FUNCTION_BLOCK "R-401_SEQ"   // FB30, GRAPH_PLUS
TITLE = Reactor R-401
{ S7_Optimized_Access := 'TRUE' }
AUTHOR : JL
VERSION : 0.1
   VAR_INPUT
      OFF_SQ : Bool := false;   // Turn sequence off
      INIT_SQ : Bool := false;   // Set sequence to initial state
      ACK_EF : Bool := false;   // Acknowledge all errors and faults
      S_PREV : Bool := false;   // Output previous step in parameter S_NO
      S_NEXT : Bool := false;   // Indicate next step in parameter S_NO
      SW_AUTO : Bool := false;   // Automatic mode
      SW_TAP : Bool := false;   // Semiautomatic/switch with transition
      SW_TOP : Bool := false;   // Semiautomatic/ignore transition
      SW_MAN : Bool := false;   // Manual mode
      S_SEL : Int := 0;   // Select step to be output to S_NO
      S_ON : Bool := false;   // Activate step indicated in S_NO
      S_OFF : Bool := false;   // Deactivate step indicated S_NO
      T_PUSH : Bool := false;   // Enable transition to switch in semi automatic mode
   END_VAR
   VAR_OUTPUT
      S_NO : Int := 0;   // Step number
      S_MORE : Bool := false;   // More steps are available and can be shown in S_NO
      S_ACTIVE : Bool := false;   // Step indicated in S_NO is active
      ERR_FLT : Bool := false;   // Interlock or supervision group error
      AUTO_ON : Bool := false;   // Automatic mode is active
      TAP_ON : Bool := false;   // Semiautomatic mode/step with transition enabled
      TOP_ON : Bool := false;   // Semiautomatic mode/ignore transition enabled
      MAN_ON : Bool := false;   // Manual mode is active
   END_VAR
   VAR
      HMI_INFO : Array[0..12] of UInt;
      IF_PAR : G7_IfParPlus_V6;
      RT_DATA : G7_RTDataPlus_V6;   // Internal data area
      Abort : G7_TransitionPlus_V6;   // Transition structure
      InitializeR : G7_TransitionPlus_V6;   // Transition structure
      CalcinP : G7_TransitionPlus_V6;   // Transition structure
      Re : G7_TransitionPlus_V6;   // Transition structure
      Calcinat : G7_TransitionPlus_V6;   // Transition structure
      Wash : G7_TransitionPlus_V6;   // Transition structure
      Shutdwn : G7_TransitionPlus_V6;   // Transition structure
      ColdDDn : G7_TransitionPlus_V6;   // Transition structure
      Std : G7_TransitionPlus_V6;   // Transition structure
      PDn : G7_TransitionPlus_V6;   // Transition structure
      PressRd : G7_TransitionPlus_V6;   // Transition structure
      Rmp1Dn : G7_TransitionPlus_V6;   // Transition structure
      FHldDn : G7_TransitionPlus_V6;   // Transition structure
      Rmp2Dn : G7_TransitionPlus_V6;   // Transition structure
      ScHldDn : G7_TransitionPlus_V6;   // Transition structure
      Rmp3Dn : G7_TransitionPlus_V6;   // Transition structure
      ThHldDn : G7_TransitionPlus_V6;   // Transition structure
      Trans30 : G7_TransitionPlus_V6;   // Transition structure
      Trans31 : G7_TransitionPlus_V6;   // Transition structure
      End : G7_TransitionPlus_V6;   // Transition structure
      Init : G7_TransitionPlus_V6;   // Transition structure
      SAut : G7_TransitionPlus_V6;   // Transition structure
      SIn : G7_TransitionPlus_V6;   // Transition structure
      Initd : G7_TransitionPlus_V6;   // Transition structure
      Ab : G7_TransitionPlus_V6;   // Transition structure
      AbortOn : G7_TransitionPlus_V6;   // Transition structure
      AbortDn : G7_TransitionPlus_V6;   // Transition structure
      ShtSted : G7_TransitionPlus_V6;   // Transition structure
      CldDwnDn : G7_TransitionPlus_V6;   // Transition structure
      DPDn : G7_TransitionPlus_V6;   // Transition structure
      Idle : G7_StepPlus_V6;   // Step structure
      Ready : G7_StepPlus_V6;   // Step structure
      SelectSeq : G7_StepPlus_V6;   // Step structure
      Started : G7_StepPlus_V6;   // Step structure
      "EDIT Params" : G7_StepPlus_V6;   // Step structure
      "USER StartAir" : G7_StepPlus_V6;   // Step structure
      RampUp1 : G7_StepPlus_V6;   // Step structure
      FirstHold : G7_StepPlus_V6;   // Step structure
      RampUp2 : G7_StepPlus_V6;   // Step structure
      SecondHold : G7_StepPlus_V6;   // Step structure
      RampUp3 : G7_StepPlus_V6;   // Step structure
      ThirdHold : G7_StepPlus_V6;   // Step structure
      HeatersOff : G7_StepPlus_V6;   // Step structure
      PressureOff : G7_StepPlus_V6;   // Step structure
      Done : G7_StepPlus_V6;   // Step structure
      Initialize : G7_StepPlus_V6;   // Step structure
      SetAuto : G7_StepPlus_V6;   // Step structure
      SetInitial : G7_StepPlus_V6;   // Step structure
      Initialized : G7_StepPlus_V6;   // Step structure
      AbortStarting : G7_StepPlus_V6;   // Step structure
      Aborting : G7_StepPlus_V6;   // Step structure
      AbortDone : G7_StepPlus_V6;   // Step structure
      ShtdnStarted : G7_StepPlus_V6;   // Step structure
      CoolingDown : G7_StepPlus_V6;   // Step structure
      DePress : G7_StepPlus_V6;   // Step structure
      ShtdnDn : G7_StepPlus_V6;   // Step structure
      SINI : Array[0..5] of USInt;
      LSTT : Array[0..29] of USInt;
      ATAJ : Array[0..29] of USInt;
      ATAB : Array[0..29] of USInt;
      PSTT : Array[0..29] of USInt;
      NSTT : Array[0..29] of USInt;
      ASSJ : Array[0..25] of USInt;
      ASSB : Array[0..25] of USInt;
      PTTS : Array[0..25] of USInt;
      NTTS : Array[0..25] of USInt;
      SW_SQTS : Array[0..25] of USInt;
      SWITCH : Array[0..4] of USInt;
      TVX : Array[0..11] of USInt;
      TTX : Array[0..11] of USInt;
      TSX : Array[0..5] of USInt;
      S00X : Array[0..5] of USInt;
      SOFFX : Array[0..5] of USInt;
      SONX : Array[0..5] of USInt;
      SAX : Array[0..5] of USInt;
      SERRX : Array[0..26] of USInt;
      SMX : Array[0..26] of USInt;
      S0X : Array[0..26] of USInt;
      S1X : Array[0..26] of USInt;
      IL_ALARM_INST : Diag_Alarm;
      SUP_ALARM_INST : Diag_Alarm;
      STEP_TIME_ALARM_INST : Diag_Alarm;
      IEC_TIMER_INST : IEC_TIMER;
      TRANSACTION_FLAG : Bool := false;
   END_VAR
   // SINI[0] := 2;
   // LSTT[0] := 19;
   // NSTT[0] := 19;
   // PTTS[0] := 255;
   // TVX[0] := 16#1;
   // TTX[0] := 16#1;
   // TSX[0] := 16#1;
   // S00X[0] := 16#1;
   // SOFFX[0] := 16#1;
   // SONX[0] := 16#1;
   // SAX[0] := 16#1;
   // SERRX[0] := 16#1;
   // SMX[0] := 16#1;
   // S0X[0] := 16#1;
   // S1X[0] := 16#1;
   // SINI[2] := 255;
   // SINI[3] := 255;
   // SINI[4] := 255;
   // LSTT[1] := 15;
   // LSTT[2] := 255;
   // LSTT[3] := 255;
   // LSTT[4] := 3;
   // LSTT[5] := 255;
   // LSTT[6] := 22;
   // LSTT[16] := 255;
   // LSTT[8] := 255;
   // LSTT[9] := 255;
   // LSTT[10] := 255;
   // LSTT[11] := 255;
   // LSTT[12] := 255;
   // LSTT[13] := 255;
   // LSTT[14] := 255;
   // LSTT[19] := 255;
   // LSTT[22] := 255;
   // LSTT[17] := 255;
   // LSTT[25] := 255;
   // LSTT[20] := 255;
   // LSTT[21] := 255;
   // ATAJ[1] := 1;
   // ATAJ[2] := 2;
   // ATAJ[3] := 3;
   // ATAJ[4] := 4;
   // ATAJ[5] := 5;
   // ATAJ[6] := 6;
   // ATAJ[7] := 7;
   // ATAJ[8] := 8;
   // ATAJ[9] := 9;
   // ATAJ[10] := 10;
   // ATAJ[11] := 11;
   // ATAJ[12] := 12;
   // ATAJ[13] := 13;
   // ATAJ[14] := 14;
   // ATAJ[15] := 15;
   // ATAJ[16] := 16;
   // ATAJ[17] := 17;
   // ATAJ[18] := 18;
   // ATAJ[19] := 19;
   // ATAJ[20] := 20;
   // ATAJ[21] := 21;
   // ATAJ[22] := 22;
   // ATAB[0] := 6;
   // ATAB[1] := 2;
   // ATAB[3] := 3;
   // ATAB[4] := 5;
   // ATAB[5] := 4;
   // ATAB[6] := 1;
   // ATAB[7] := 7;
   // ATAB[8] := 8;
   // ATAB[9] := 9;
   // ATAB[10] := 10;
   // ATAB[11] := 11;
   // ATAB[12] := 12;
   // ATAB[13] := 13;
   // ATAB[14] := 14;
   // ATAB[15] := 15;
   // ATAB[16] := 16;
   // ATAB[17] := 17;
   // ATAB[18] := 18;
   // ATAB[19] := 19;
   // ATAB[20] := 20;
   // ATAB[21] := 21;
   // ATAB[22] := 22;
   // SW_SQTS[21] := 4;
   // SW_SQTS[20] := 4;
   // PSTT[3] := 1;
   // PSTT[4] := 2;
   // PSTT[5] := 2;
   // PSTT[22] := 17;
   // PSTT[7] := 25;
   // PSTT[8] := 3;
   // PSTT[9] := 4;
   // PSTT[10] := 5;
   // PSTT[11] := 6;
   // PSTT[12] := 7;
   // PSTT[13] := 8;
   // PSTT[14] := 9;
   // PSTT[15] := 10;
   // PSTT[16] := 11;
   // PSTT[17] := 13;
   // PSTT[18] := 14;
   // PSTT[19] := 12;
   // PSTT[20] := 15;
   // PSTT[21] := 16;
   // PSTT[25] := 20;
   // NTTS[21] := 26;
   // NTTS[20] := 25;
   // PTTS[21] := 25;
   // PTTS[20] := 24;
   // NSTT[1] := 15;
   // NSTT[2] := 1;
   // NSTT[3] := 2;
   // NSTT[4] := 3;
   // NSTT[5] := 255;
   // NSTT[6] := 22;
   // NSTT[16] := 12;
   // NSTT[8] := 4;
   // NSTT[9] := 5;
   // NSTT[10] := 6;
   // NSTT[11] := 7;
   // NSTT[12] := 8;
   // NSTT[13] := 9;
   // NSTT[14] := 10;
   // NSTT[19] := 13;
   // NSTT[22] := 18;
   // NSTT[17] := 14;
   // NSTT[25] := 21;
   // NSTT[20] := 16;
   // NSTT[21] := 17;
   // ASSJ[20] := 20;
   // ASSB[21] := 21;
   // ASSB[20] := 20;
   // ASSJ[21] := 21;
   // ASSJ[1] := 1;
   // ASSJ[2] := 2;
   // ASSJ[3] := 3;
   // ASSJ[4] := 4;
   // ASSJ[5] := 5;
   // ASSJ[6] := 6;
   // ASSJ[7] := 7;
   // ASSJ[8] := 8;
   // ASSJ[9] := 9;
   // ASSJ[10] := 10;
   // ASSJ[11] := 11;
   // ASSJ[12] := 12;
   // ASSJ[13] := 13;
   // ASSJ[14] := 14;
   // ASSJ[15] := 15;
   // ASSJ[16] := 16;
   // ASSJ[17] := 17;
   // ASSJ[18] := 18;
   // ASSJ[19] := 19;
   // NSTT[23] := 1;
   // NSTT[15] := 11;
   // PSTT[24] := 19;
   // PSTT[23] := 18;
   // ASSB[1] := 1;
   // ASSB[2] := 2;
   // ASSB[3] := 3;
   // ASSB[4] := 4;
   // ASSB[5] := 5;
   // ASSB[6] := 6;
   // ASSB[7] := 7;
   // ASSB[8] := 8;
   // ASSB[9] := 9;
   // ASSB[10] := 10;
   // ASSB[11] := 11;
   // ASSB[12] := 12;
   // ASSB[13] := 13;
   // ASSB[14] := 14;
   // ASSB[15] := 15;
   // ASSB[16] := 16;
   // ASSB[17] := 17;
   // ASSB[18] := 18;
   // ASSB[19] := 19;
   // ATAB[24] := 24;
   // ATAB[23] := 23;
   // ATAJ[24] := 24;
   // ATAJ[23] := 23;
   // PTTS[1] := 2;
   // PTTS[2] := 3;
   // PTTS[3] := 255;
   // PTTS[4] := 8;
   // PTTS[5] := 9;
   // PTTS[6] := 10;
   // PTTS[7] := 11;
   // PTTS[8] := 12;
   // PTTS[9] := 13;
   // PTTS[10] := 14;
   // PTTS[11] := 15;
   // PTTS[12] := 16;
   // PTTS[13] := 19;
   // PTTS[14] := 17;
   // PTTS[15] := 255;
   // PTTS[16] := 20;
   // PTTS[17] := 21;
   // PTTS[18] := 22;
   // PTTS[19] := 255;
   // LSTT[23] := 1;
   // LSTT[15] := 255;
   // NTTS[1] := 3;
   // NTTS[2] := 4;
   // NTTS[3] := 8;
   // NTTS[4] := 9;
   // NTTS[5] := 10;
   // NTTS[6] := 11;
   // NTTS[7] := 12;
   // NTTS[8] := 13;
   // NTTS[9] := 14;
   // NTTS[10] := 15;
   // NTTS[11] := 16;
   // NTTS[12] := 19;
   // NTTS[13] := 17;
   // NTTS[14] := 18;
   // NTTS[15] := 20;
   // NTTS[16] := 21;
   // NTTS[17] := 22;
   // NTTS[18] := 23;
   // NTTS[19] := 24;
   // SW_SQTS[1] := 1;
   // SW_SQTS[2] := 1;
   // SW_SQTS[3] := 2;
   // SW_SQTS[4] := 2;
   // SW_SQTS[5] := 2;
   // SW_SQTS[6] := 2;
   // SW_SQTS[7] := 2;
   // SW_SQTS[8] := 2;
   // SW_SQTS[9] := 2;
   // SW_SQTS[10] := 2;
   // SW_SQTS[11] := 2;
   // SW_SQTS[12] := 2;
   // SW_SQTS[13] := 2;
   // SW_SQTS[14] := 2;
   // SW_SQTS[15] := 3;
   // SW_SQTS[16] := 3;
   // SW_SQTS[17] := 3;
   // SW_SQTS[18] := 3;
   // SW_SQTS[19] := 4;
   // SWITCH[0] := 60;
   // SWITCH[1] := 191;
   // SWITCH[2] := 223;
   // SINI[5] := 255;
   // LSTT[24] := 255;
   // LSTT[28] := 255;
   // LSTT[27] := 255;
   // ATAJ[25] := 25;
   // ATAJ[26] := 26;
   // ATAJ[27] := 27;
   // ATAJ[28] := 28;
   // ATAB[25] := 25;
   // ATAB[26] := 26;
   // ATAB[27] := 27;
   // ATAB[28] := 28;
   // PSTT[26] := 21;
   // PSTT[27] := 22;
   // PSTT[28] := 23;
   // NSTT[24] := 20;
   // NSTT[28] := 24;
   // NSTT[27] := 23;
   // ASSJ[22] := 22;
   // ASSJ[23] := 23;
   // ASSJ[24] := 24;
   // ASSB[22] := 22;
   // ASSB[23] := 23;
   // ASSB[24] := 24;
   // PTTS[22] := 255;
   // PTTS[23] := 27;
   // PTTS[24] := 28;
   // NTTS[22] := 27;
   // NTTS[23] := 28;
   // NTTS[24] := 29;
   // SW_SQTS[22] := 5;
   // SW_SQTS[23] := 5;
   // SW_SQTS[24] := 5;
   // SWITCH[3] := 239;
   // SWITCH[4] := 7;
   // LSTT[29] := 255;
   // ATAJ[29] := 29;
   // ATAB[29] := 29;
   // PSTT[29] := 24;
   // NSTT[29] := 25;
   // ASSJ[25] := 25;
   // ASSB[25] := 25;
   // PTTS[25] := 29;
   // NTTS[25] := 7;
   // SW_SQTS[25] := 5;
BEGIN
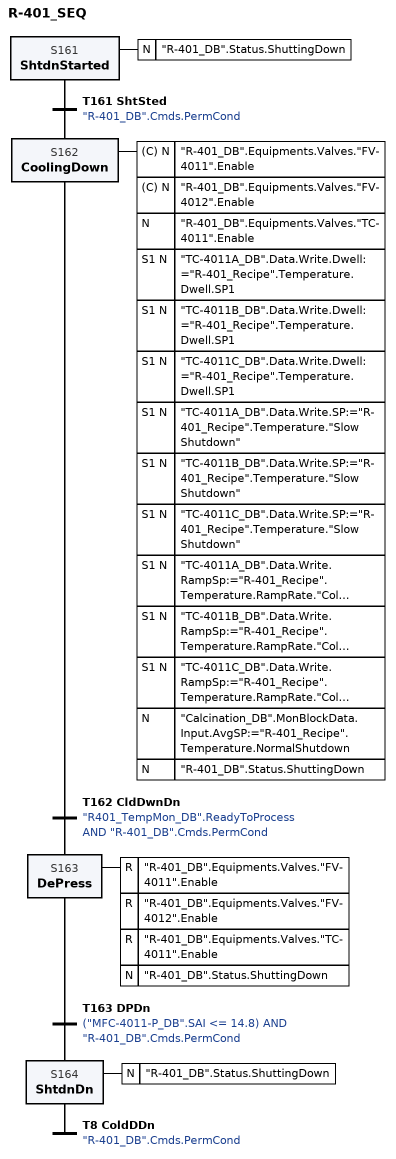
   // permanent pre-instructions
   NETWORK 1
      "R-401_SEQ_FC"();
      "R-401_FC_Inputs"();
      "Monitor_SEQ_FC"();
      "R-401_Tansitions_FC"();
      "Alarms"();

   // sequencer 1
   STEP ShtdnStarted:   // S161, max time T#10S, warning time T#7S
      // Shutdown Started
              N    "R-401_DB".Status.ShuttingDown
   END_STEP
   TRANSITION ShtSted FROM ShtdnStarted TO CoolingDown   // T161
      := "R-401_DB".Cmds.PermCond;
   END_TRANSITION
   STEP CoolingDown:   // S162, max time T#10S, warning time T#7S
      interlock C := "R-401_DB".Cmds.IL;
      (C)     N    "R-401_DB".Equipments.Valves."FV-4011".Enable
      (C)     N    "R-401_DB".Equipments.Valves."FV-4012".Enable
              N    "R-401_DB".Equipments.Valves."TC-4011".Enable
          S1  N    "TC-4011A_DB".Data.Write.Dwell:="R-401_Recipe".Temperature.Dwell.SP1
          S1  N    "TC-4011B_DB".Data.Write.Dwell:="R-401_Recipe".Temperature.Dwell.SP1
          S1  N    "TC-4011C_DB".Data.Write.Dwell:="R-401_Recipe".Temperature.Dwell.SP1
          S1  N    "TC-4011A_DB".Data.Write.SP:="R-401_Recipe".Temperature."Slow Shutdown"
          S1  N    "TC-4011B_DB".Data.Write.SP:="R-401_Recipe".Temperature."Slow Shutdown"
          S1  N    "TC-4011C_DB".Data.Write.SP:="R-401_Recipe".Temperature."Slow Shutdown"
          S1  N    "TC-4011A_DB".Data.Write.RampSp:="R-401_Recipe".Temperature.RampRate."Cold Down"
          S1  N    "TC-4011B_DB".Data.Write.RampSp:="R-401_Recipe".Temperature.RampRate."Cold Down"
          S1  N    "TC-4011C_DB".Data.Write.RampSp:="R-401_Recipe".Temperature.RampRate."Cold Down"
              N    "Calcination_DB".MonBlockData.Input.AvgSP:="R-401_Recipe".Temperature.NormalShutdown
              N    "R-401_DB".Status.ShuttingDown
   END_STEP
   TRANSITION CldDwnDn FROM CoolingDown TO DePress   // T162
      := "R401_TempMon_DB".ReadyToProcess AND "R-401_DB".Cmds.PermCond;
   END_TRANSITION
   STEP DePress:   // S163, max time T#10S, warning time T#7S
              R    "R-401_DB".Equipments.Valves."FV-4011".Enable
              R    "R-401_DB".Equipments.Valves."FV-4012".Enable
              R    "R-401_DB".Equipments.Valves."TC-4011".Enable
              N    "R-401_DB".Status.ShuttingDown
   END_STEP
   TRANSITION DPDn FROM DePress TO ShtdnDn   // T163
      := ("MFC-4011-P_DB".SAI <= 14.8) AND "R-401_DB".Cmds.PermCond;
   END_TRANSITION
   STEP ShtdnDn:   // S164, max time T#10S, warning time T#7S
              N    "R-401_DB".Status.ShuttingDown
   END_STEP
   TRANSITION ColdDDn FROM ShtdnDn TO ?   // T8
      := "R-401_DB".Cmds.PermCond;
   END_TRANSITION

   // permanent post-instructions
   NETWORK 1
      "R-401_FC_Outputs"();
END_FUNCTION_BLOCK

FUNCTION "R-401_FC_Inputs" : Void   // FC51, SCL
{ S7_Optimized_Access := 'TRUE' }
VERSION : 0.1
   VAR_TEMP
      fdfdfd : DInt;
   END_VAR
BEGIN
   //************************************************************************************************************************************
   //************************************************From Eurotherm TC-401A Controllers*********************************************************
   //***************************************************** Working Setpoint (SP)********************************************************

   IF "R-402_Aux_DB"."Bool".EurothermStatus."4011A_Connected" THEN     //Check if Modbus Connection is Ok
       "TC-4011A_DB".Data.Read.WorkingSP := INT_TO_REAL("TC-4011A_R1".MB_Data.Buffer[5]);
   ELSE
       "TC-4011A_DB".Data.Read.WorkingSP := 0.0;
   END_IF;

   IF "R-402_Aux_DB"."Bool".EurothermStatus."4011B_Connected" THEN     //Check if Modbus Connection is Ok
       "TC-4011B_DB".Data.Read.WorkingSP := INT_TO_REAL("TC-4011B_R1".MB_Data.Buffer[5]);
   ELSE
       "TC-4011B_DB".Data.Read.WorkingSP := 0.0;
   END_IF;

   IF "R-402_Aux_DB"."Bool".EurothermStatus."4011C_Connected" THEN     //Check if Modbus Connection is Ok
       "TC-4011C_DB".Data.Read.WorkingSP := INT_TO_REAL("TC-4011C_R1".MB_Data.Buffer[5]);
   ELSE
       "TC-4011C_DB".Data.Read.WorkingSP := 0.0;
   END_IF;

   //*****************************************************Process Value (PV)********************************************************

   IF "R-402_Aux_DB"."Bool".EurothermStatus."4011A_Connected" THEN     //Check if Modbus Connection is Ok
       "TC-4011A_DB".Data.Read.PV := INT_TO_REAL("TC-4011A_R1".MB_Data.Buffer[1]);
   ELSE
       "TC-4011A_DB".Data.Read.PV := 0.0;
   END_IF;

   IF "R-402_Aux_DB"."Bool".EurothermStatus."4011B_Connected" THEN     //Check if Modbus Connection is Ok
       "TC-4011B_DB".Data.Read.PV := INT_TO_REAL("TC-4011B_R1".MB_Data.Buffer[1]);
   ELSE
       "TC-4011B_DB".Data.Read.PV := 0.0;
   END_IF;

   IF "R-402_Aux_DB"."Bool".EurothermStatus."4011C_Connected" THEN     //Check if Modbus Connection is Ok
       "TC-4011C_DB".Data.Read.PV := INT_TO_REAL("TC-4011C_R1".MB_Data.Buffer[1]);
   ELSE
       "TC-4011C_DB".Data.Read.PV := 0.0;
   END_IF;


   //***************************************************** Controller Output (OP)******************************************************

   IF "R-402_Aux_DB"."Bool".EurothermStatus."4011A_Connected" THEN     //Check if Modbus Connection is Ok
       "TC-4011A_DB".Data.Read.OP := INT_TO_REAL("TC-4011A_R1".MB_Data.Buffer[4]/10);
   ELSE
       "TC-4011A_DB".Data.Read.OP := 0.0;
   END_IF;

   IF "R-402_Aux_DB"."Bool".EurothermStatus."4011B_Connected" THEN     //Check if Modbus Connection is Ok
       "TC-4011B_DB".Data.Read.OP := INT_TO_REAL("TC-4011B_R1".MB_Data.Buffer[4] / 10);
   ELSE
       "TC-4011B_DB".Data.Read.OP := 0.0;
   END_IF;

   IF "R-402_Aux_DB"."Bool".EurothermStatus."4011C_Connected" THEN     //Check if Modbus Connection is Ok
       "TC-4011C_DB".Data.Read.OP := INT_TO_REAL("TC-4011C_R1".MB_Data.Buffer[4]/10);
   ELSE
       "TC-4011C_DB".Data.Read.OP := 0.0;
   END_IF;
END_FUNCTION

FUNCTION "R-401_FC_Outputs" : Void   // FC85, SCL
{ S7_Optimized_Access := 'TRUE' }
VERSION : 0.1
   VAR_TEMP
      "FV-4011" : Struct
         On : Bool;
         Cond_1 : Bool;
      END_STRUCT;
      "FV-4012" : Struct
         On : Bool;
         Cond_1 : Bool;
      END_STRUCT;
      "TC-4011" : Struct
         On : Bool;
         Cond_1 : Bool;
      END_STRUCT;
   END_VAR
BEGIN
   //****** Equipmens Activation*******
   //**********************************TC-4011 Eurotherm Temperature Control (TC-4011)**************************************************

   #"TC-4011".Cond_1 := "R-401_DB".Equipments.Valves."TC-4011".Enable AND NOT "R-401_Aux_DB".Timer.HoldTimer.Q;
       "R-401_DB".Equipments.Valves."TC-4011".CmdOn := #"TC-4011".Cond_1 AND NOT "R-401_DB".Cmds.Hold AND NOT "R-401_DB".Status.Aborting;
       //Delay Off 
       #"TC-4011".On := "R-401_DB".Equipments.Valves."TC-4011".CmdOn;

       IF #"TC-4011".On AND ("R-401_DB".Status.Step=24 OR "R-401_DB".Status.Step=26 OR "R-401_DB".Status.Step=28) AND "R-401_Aux_DB"."Bool".Cond._005 THEN //Run Command for the Eurotherm Controllers
           "TC-4011A_DB".Data.Write.CMD := 1;
           "TC-4011B_DB".Data.Write.CMD  := 1;
           "TC-4011C_DB".Data.Write.CMD  := 1;

           //**********Working SP Reached ********
           "R-401_Aux_DB"."Bool".Cond._006 := "TC-4011A_DB".Data.Write.SP = "TC-4011A_DB".Data.Read.WorkingSP;
           "R-401_Aux_DB"."Bool".Cond._007 := "TC-4011B_DB".Data.Write.SP = "TC-4011B_DB".Data.Read.WorkingSP;
           "R-401_Aux_DB"."Bool".Cond._008 := "TC-4011C_DB".Data.Write.SP = "TC-4011C_DB".Data.Read.WorkingSP;

           "R-401_Aux_DB"."Bool".Cond._009 := "R-401_Aux_DB"."Bool".Cond._006 AND "R-401_Aux_DB"."Bool".Cond._007 AND "R-401_Aux_DB"."Bool".Cond._008;

       ELSIF #"TC-4011".On AND ("R-401_DB".Status.Step=25 OR "R-401_DB".Status.Step=27 OR "R-401_DB".Status.Step=29) AND "R-401_Aux_DB"."Bool".Cond._005 THEN //Hold command for the Eurotherm Controllers
           "TC-4011A_DB".Data.Write.CMD  := 2;
           "TC-4011B_DB".Data.Write.CMD  := 2;
           "TC-4011C_DB".Data.Write.CMD  := 2;

           "R-401_Aux_DB"."Bool".Cond._009 := FALSE;
       ELSE    //Stop Command for the Eurotherm Controllers
           "TC-4011A_DB".Data.Write.CMD  := 0;
           "TC-4011B_DB".Data.Write.CMD  := 0;
           "TC-4011C_DB".Data.Write.CMD  := 0;

           "R-401_Aux_DB"."Bool".Cond._009 := FALSE;
       END_IF;
       "R-401_DB".Equipments.Valves."TC-4011".TurningOff := NOT "R-401_DB".Equipments.Valves."TC-4011".CmdOn AND "R-401_Aux_DB".Timer."TC-4011".Q;

   //**********************************FV-4011 Air Pressure Control Valve (MFC-4011)******************************************************
   IF "FV-4011_DB".HMI.Config.Mode = 0 THEN
       #"FV-4011".Cond_1 := "R-401_DB".Equipments.Valves."FV-4011".Enable;
       "R-401_DB".Equipments.Valves."FV-4011".CmdOn := #"FV-4011".Cond_1 AND NOT "R-401_DB".Cmds.Hold AND NOT "R-401_DB".Status.Aborting;
       //Delay Off To avoid Overpressure the Lines
       #"FV-4011".On := "R-401_DB".Equipments.Valves."FV-4011".CmdOn;
       "R-401_Aux_DB".Timer."FV-4011".TOF(IN := #"FV-4011".On,
                                          PT := "R-401_Aux_DB".Constants.CmdDelay);
       IF "R-401_Aux_DB".Timer."FV-4011".Q  THEN

           // "MFC-4011_DB_MB".Data.SP := "R-401_Recipe".Pressure.Calcination;

           "MFC-4011_DB".enableManualMode := False;
           "MFC-4011_DB".enableRemoteSetpoint := False;
            "MFC-4011_DB".hmi.Controls.manualEnable := False;
            "MFC-4011_DB".hmi.Config.mode := 3;

       END_IF;
      // ELSE
          // "MFC-4011_DB".enableManualMode := True;
          // "MFC-4011_DB".hmi.Controls.manualEnable := True;
          // "MFC-4011_DB".hmi.Config.mode := 4;
          // "MFC-4011_DB".hmi.Controls.manualOutput := "R-401_Recipe".Pressure.Shutdown;

          // "MFC-4011_DB_MB".Data.SP := "R-401_Recipe".Pressure.Shutdown;

      // END_IF;
       "R-401_DB".Equipments.Valves."FV-4011".TurningOff := NOT "R-401_DB".Equipments.Valves."FV-4011".CmdOn AND "R-401_Aux_DB".Timer."FV-4011".Q;
   END_IF;

   //**********************************FV-4012 N2 Pressure Control Valve (MFC-4012)******************************************************
   IF "FV-4012_DB".HMI.Config.Mode = 0 THEN
       #"FV-4012".Cond_1 := "R-401_DB".Equipments.Valves."FV-4012".Enable;
       "R-401_DB".Equipments.Valves."FV-4012".CmdOn := #"FV-4012".Cond_1 AND NOT "R-401_DB".Cmds.Hold AND NOT "R-401_DB".Status.Aborting;
       //Delay Off To avoid Overpressure the Lines
       #"FV-4012".On := "R-401_DB".Equipments.Valves."FV-4012".CmdOn;
       "R-401_Aux_DB".Timer."FV-4012".TOF(IN := #"FV-4012".On,
                                          PT := "R-401_Aux_DB".Constants.CmdDelay);
       IF "R-401_Aux_DB".Timer."FV-4012".Q THEN

           // "MFC-4011_DB_MB".Data.SP := "R-401_Recipe".Pressure.Calcination;

           "MFC-4012_DB".enableManualMode := False;
           "MFC-4012_DB".enableRemoteSetpoint := False;
           "MFC-4012_DB".hmi.Controls.manualEnable := False;
           "MFC-4012_DB".hmi.Config.mode := 3;

       END_IF;
       // ELSE
       // "MFC-4011_DB".enableManualMode := True;
       // "MFC-4011_DB".hmi.Controls.manualEnable := True;
       // "MFC-4011_DB".hmi.Config.mode := 4;
       // "MFC-4011_DB".hmi.Controls.manualOutput := "R-401_Recipe".Pressure.Shutdown;

       // "MFC-4011_DB_MB".Data.SP := "R-401_Recipe".Pressure.Shutdown;

       // END_IF;
       "R-401_DB".Equipments.Valves."FV-4012".TurningOff := NOT "R-401_DB".Equipments.Valves."FV-4012".CmdOn AND "R-401_Aux_DB".Timer."FV-4012".Q;
   END_IF;
   //******************************************************************************************************************************************//
   //**************************************************To Temperature Controllers**************************************************************

       //***********************************************Temperature Controllers Commands*******************************************************//
   "TC-4011A_W1".MB_Data.Buffer[1] := "TC-4011A_DB".Data.Write.CMD;
   "TC-4011B_W1".MB_Data.Buffer[1]:= "TC-4011B_DB".Data.Write.CMD;
   "TC-4011C_W1".MB_Data.Buffer[1] := "TC-4011C_DB".Data.Write.CMD;

   //***********************************************Dwell to Temperature Controllers ******************************************************//
   IF "TC-4011A_DB".Data.Write.Dwell = "TC-4011A_R2".MB_Data.Buffer[1]
       AND "TC-4011A_DB".Data.Write.Dwell = "TC-4011B_R2".MB_Data.Buffer[1]
       AND "TC-4011A_DB".Data.Write.Dwell = "TC-4011C_R2".MB_Data.Buffer[1] THEN    //Compare read value and SP to activate or deactivate the Modbus Write block

       "TC-4011A_W2".Disconnect := TRUE;
       "TC-4011B_W2".Disconnect := TRUE;
       "TC-4011C_W2".Disconnect := TRUE;
       "R-401_Aux_DB"."Bool".Cond._004 := TRUE;
   ELSE
       "TC-4011A_W2".MB_Data.Buffer[1] := "TC-4011A_DB".Data.Write.Dwell;
       "TC-4011B_W2".MB_Data.Buffer[1] := "TC-4011B_DB".Data.Write.Dwell;
       "TC-4011C_W2".MB_Data.Buffer[1] := "TC-4011C_DB".Data.Write.Dwell;
       "TC-4011A_W2".Disconnect := FALSE;
       "TC-4011B_W2".Disconnect := FALSE;
       "TC-4011C_W2".Disconnect := FALSE;
       "R-401_Aux_DB"."Bool".Cond._004 := FALSE;
   END_IF;
       //***********************************************Temperature Controllers SetPoints*****************************************************//
   IF "TC-4011A_DB".Data.Write.SP = "TC-4011A_R2".MB_Data.Buffer[2]    
       AND "TC-4011A_DB".Data.Write.SP = "TC-4011B_R2".MB_Data.Buffer[2]
       AND "TC-4011A_DB".Data.Write.SP = "TC-4011C_R2".MB_Data.Buffer[2] THEN   //Compare read value and SP to activate or deactivate the Modbus Write block
       "TC-4011A_W3".Disconnect := TRUE;
       "TC-4011B_W3".Disconnect := TRUE;
       "TC-4011C_W3".Disconnect := TRUE;
       "R-401_Aux_DB"."Bool".Cond._002 := TRUE;        //Temperature SP
   ELSE
       "TC-4011A_W3".MB_Data.Buffer[1] := REAL_TO_INT("TC-4011A_DB".Data.Write.SP);
       "TC-4011B_W3".MB_Data.Buffer[1] := REAL_TO_INT("TC-4011B_DB".Data.Write.SP);
       "TC-4011C_W3".MB_Data.Buffer[1] := REAL_TO_INT("TC-4011C_DB".Data.Write.SP);
       "TC-4011A_W3".Disconnect := FALSE;
       "TC-4011B_W3".Disconnect := FALSE;
       "TC-4011C_W3".Disconnect := FALSE;
       "R-401_Aux_DB"."Bool".Cond._002 := FALSE;       //Temperature SP
   END_IF;
       //***********************************************Temperature Controllers Ramp Rate SetPoints*******************************************//
   IF "TC-4011A_DB".Data.Write.RampSp = "TC-4011A_R2".MB_Data.Buffer[3]/10
       AND "TC-4011A_DB".Data.Write.RampSp = "TC-4011B_R2".MB_Data.Buffer[3]/10
       AND "TC-4011A_DB".Data.Write.RampSp = "TC-4011C_R2".MB_Data.Buffer[3]/10 THEN   //Compare read value and SP to activate or deactivate the Modbus Write block

       "TC-4011A_W4".Disconnect := TRUE;
       "TC-4011B_W4".Disconnect := TRUE;
       "TC-4011C_W4".Disconnect := TRUE;
       "R-401_Aux_DB"."Bool".Cond._003 := TRUE;
   ELSE
       "TC-4011A_W4".MB_Data.Buffer[1] := "TC-4011A_DB".Data.Write.RampSp*10;
       "TC-4011B_W4".MB_Data.Buffer[1] := "TC-4011B_DB".Data.Write.RampSp*10;
       "TC-4011C_W4".MB_Data.Buffer[1] := "TC-4011C_DB".Data.Write.RampSp*10;
       "TC-4011A_W4".Disconnect := FALSE;
       "TC-4011B_W4".Disconnect := FALSE;
       "TC-4011C_W4".Disconnect := FALSE;
       "R-401_Aux_DB"."Bool".Cond._003 := FALSE;
   END_IF;

   "R-401_Aux_DB"."Bool".Cond._005 := "R-401_Aux_DB"."Bool".Cond._002 AND "R-401_Aux_DB"."Bool".Cond._003 AND "R-401_Aux_DB"."Bool".Cond._004;

   //**********ALICAT Controllers************//
       //***********************************************ALICAT Control Selection*******************************************************//
       //Command ID and Command Argument 
       (*With this Values the Selection is:
           Address 1000=11; Change control loop variable
           Address 1001=3;  Absolute Pressure*)
       //*********MFC-4011*********
       "MFC-4011_MB_WCMD_DB".MB_Data.Buffer[1] := 11;
       "MFC-4011_MB_WCMD_DB".MB_Data.Buffer[2] := 3;
       //*********MFC-4012*********
       "MFC-4012_MB_WCMD_DB".MB_Data.Buffer[1] := 11;
       "MFC-4012_MB_WCMD_DB".MB_Data.Buffer[2] := 3;
       //***********************************************ALICAT Controller Set Point*******************************************************//
       //*********MFC-4011*********
       "MFC-4011_MB_W_DB".MB_Data.Buffer[1] := (INT_TO_REAL("FV-4011_DB".CMD) * 100) / 27648.0;
       "MFC-4011_DB_MB".Data.SP := "MFC-4011_MB_W_DB".MB_Data.Buffer[1];
       //*********MFC-4012*********
       "MFC-4012_MB_W_DB".MB_Data.Buffer[1] := (INT_TO_REAL("FV-4012_DB".CMD) * 100) / 27648.0;
       "MFC-4012_DB_MB".Data.SP := "MFC-4012_MB_W_DB".MB_Data.Buffer[1];

       //***************************************************Setpoints Ranges***************************************************************
       IF "R-401_DB".Status.Step = 24 OR "R-401_DB".Status.Step = 25 THEN
           "Calcination_DB".MonBlockData.Input."Min Range" := "R-401_Recipe".Temperature.SP1 - "R-401_Aux_DB"."Real"."TE-401".Temperature.MinRange;
           "Calcination_DB".MonBlockData.Input."Max Range" := "R-401_Recipe".Temperature.SP1 + "R-401_Aux_DB"."Real"."TE-401".Temperature.MaxRange;
       ELSIF "R-401_DB".Status.Step = 26 OR "R-401_DB".Status.Step = 27 THEN
           "Calcination_DB".MonBlockData.Input."Min Range" := "R-401_Recipe".Temperature.SP2 - "R-401_Aux_DB"."Real"."TE-401".Temperature.MinRange;
           "Calcination_DB".MonBlockData.Input."Max Range" := "R-401_Recipe".Temperature.SP2 + "R-401_Aux_DB"."Real"."TE-401".Temperature.MaxRange;
       ELSIF "R-401_DB".Status.Step = 28 OR "R-401_DB".Status.Step = 29  THEN
           "Calcination_DB".MonBlockData.Input."Min Range" := "R-401_Recipe".Temperature.SP3 - "R-401_Aux_DB"."Real"."TE-401".Temperature.MinRange;
           "Calcination_DB".MonBlockData.Input."Max Range" := "R-401_Recipe".Temperature.SP3 + "R-401_Aux_DB"."Real"."TE-401".Temperature.MaxRange;
       END_IF;

       "Calcination_DB".MonBlockData.Input.MinAvgValue := "R-401_Aux_DB"."Real"."TE-401".Temperature.MinAvgValue;
       "Calcination_DB".MonBlockData.Input.MaxAvgValue := "R-401_Aux_DB"."Real"."TE-401".Temperature.MaxAvgValue;
       "Calcination_DB".MonBlockData.Input.AlarmDeviation := "R-401_Aux_DB"."Real"."TE-401".Temperature.AlarmDeviation;
       "Calcination_DB".MonBlockData.Input.MaxDeviation := "R-401_Aux_DB"."Real"."TE-401".Temperature.MaxDeviation;



       //***************Valves Status***************//
       "R-401_Aux_DB"."Bool".TOff := "R-401_DB".Equipments.Valves."FV-4011".TurningOff;

       //***********************************************Timers****************************************************************************//
       "R-401_Aux_DB"."Bool".HoldTimeEn := ("R-401_SEQ_DB".S_NO = 25 OR "R-401_SEQ_DB".S_NO = 27 OR "R-401_SEQ_DB".S_NO = 29); //"R401_TempMon_DB".ReadyToProcess AND 
       "R-401_Aux_DB"."Bool".HoldTime_Reset := "R-401_DB".Status.Step = 1 OR (NOT "R401_TempMon_DB".ReadyToProcess AND ("R-401_SEQ_DB".S_NO = 24 OR "R-401_SEQ_DB".S_NO = 26 OR "R-401_SEQ_DB".S_NO = 28 OR "R-401_SEQ_DB".S_NO = 30));
END_FUNCTION

FUNCTION "R-401_SEQ_FC" : Void   // FC92, LAD
{ S7_Optimized_Access := 'TRUE' }
VERSION : 0.1
   VAR_TEMP   // added for the SCL form of the ladder/FBD networks
      _w1 : Bool;
      _w2 : Bool;
      _w3 : Bool;
   END_VAR
BEGIN

REGION Network 2: Abort/Shutdown
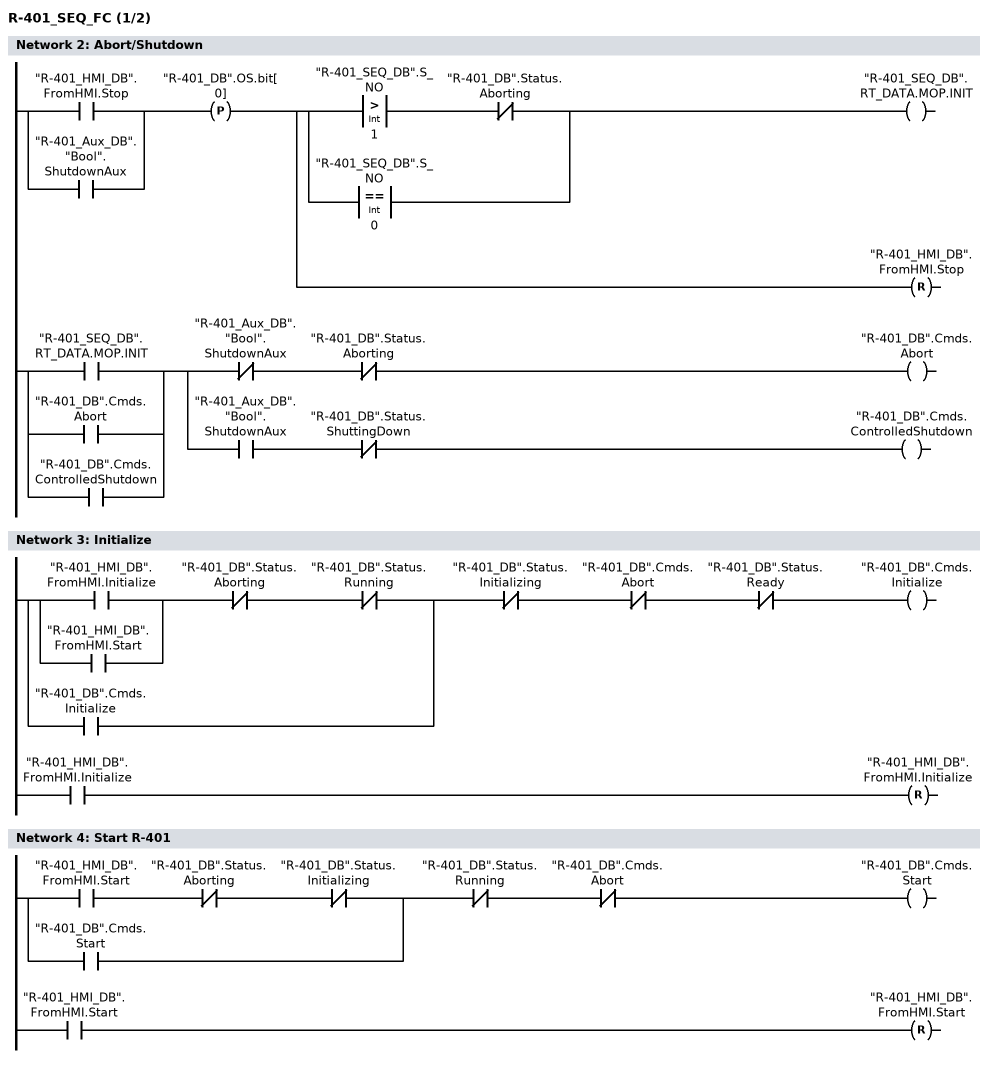
   RUNG wire#powerrail
      Contact( "R-401_HMI_DB".FromHMI.Stop )
      wire#w1
      P_Trig( "R-401_DB".OS.bit[0] )
      wire#w2
      { S7_Templates := "SrcType := Int" } GT_Contact(in1 := "R-401_SEQ_DB".S_NO, in2 := 1)
      I_Contact( "R-401_DB".Status.Aborting )
      wire#w3
      Coil( "R-401_SEQ_DB".RT_DATA.MOP.INIT )
   END_RUNG
   RUNG wire#powerrail
      Contact( "R-401_Aux_DB"."Bool".ShutdownAux )
   END_RUNG wire#w1
   RUNG wire#w2
      { S7_Templates := "SrcType := Int" } EQ_Contact(in1 := "R-401_SEQ_DB".S_NO, in2 := 0)
   END_RUNG wire#w3
   RUNG wire#w2
      R_Coil( "R-401_HMI_DB".FromHMI.Stop )
   END_RUNG
   RUNG wire#powerrail
      Contact( "R-401_SEQ_DB".RT_DATA.MOP.INIT )
      wire#w4
      I_Contact( "R-401_Aux_DB"."Bool".ShutdownAux )
      I_Contact( "R-401_DB".Status.Aborting )
      Coil( "R-401_DB".Cmds.Abort )
   END_RUNG
   RUNG wire#powerrail
      Contact( "R-401_DB".Cmds.Abort )
   END_RUNG wire#w4
   RUNG wire#powerrail
      Contact( "R-401_DB".Cmds.ControlledShutdown )
   END_RUNG wire#w4
   RUNG wire#w4
      Contact( "R-401_Aux_DB"."Bool".ShutdownAux )
      I_Contact( "R-401_DB".Status.ShuttingDown )
      Coil( "R-401_DB".Cmds.ControlledShutdown )
   END_RUNG
   // the same network as SCL:
   #_w1 := "R-401_HMI_DB".FromHMI.Stop OR "R-401_Aux_DB"."Bool".ShutdownAux;
   #_w2 := #_w1 AND NOT "R-401_DB".OS.bit[0];   // rising edge
   "R-401_DB".OS.bit[0] := #_w1;
   "R-401_SEQ_DB".RT_DATA.MOP.INIT := #_w2 AND ((("R-401_SEQ_DB".S_NO > 1) AND NOT "R-401_DB".Status.Aborting) OR ("R-401_SEQ_DB".S_NO = 0));
   IF #_w2 THEN "R-401_HMI_DB".FromHMI.Stop := FALSE; END_IF;
   #_w3 := "R-401_SEQ_DB".RT_DATA.MOP.INIT OR "R-401_DB".Cmds.Abort OR "R-401_DB".Cmds.ControlledShutdown;
   "R-401_DB".Cmds.Abort := #_w3 AND NOT "R-401_Aux_DB"."Bool".ShutdownAux AND NOT "R-401_DB".Status.Aborting;
   "R-401_DB".Cmds.ControlledShutdown := #_w3 AND "R-401_Aux_DB"."Bool".ShutdownAux AND NOT "R-401_DB".Status.ShuttingDown;
END_REGION

REGION Network 3: Initialize
   RUNG wire#powerrail
      Contact( "R-401_HMI_DB".FromHMI.Initialize )
      wire#w1
      I_Contact( "R-401_DB".Status.Aborting )
      I_Contact( "R-401_DB".Status.Running )
      wire#w2
      I_Contact( "R-401_DB".Status.Initializing )
      I_Contact( "R-401_DB".Cmds.Abort )
      I_Contact( "R-401_DB".Status.Ready )
      Coil( "R-401_DB".Cmds.Initialize )
   END_RUNG
   RUNG wire#powerrail
      Contact( "R-401_HMI_DB".FromHMI.Start )
   END_RUNG wire#w1
   RUNG wire#powerrail
      Contact( "R-401_DB".Cmds.Initialize )
   END_RUNG wire#w2
   RUNG wire#powerrail
      Contact( "R-401_HMI_DB".FromHMI.Initialize )
      R_Coil( "R-401_HMI_DB".FromHMI.Initialize )
   END_RUNG
   // the same network as SCL:
   "R-401_DB".Cmds.Initialize := ((("R-401_HMI_DB".FromHMI.Initialize OR "R-401_HMI_DB".FromHMI.Start) AND NOT "R-401_DB".Status.Aborting AND NOT "R-401_DB".Status.Running) OR "R-401_DB".Cmds.Initialize) AND NOT "R-401_DB".Status.Initializing AND NOT "R-401_DB".Cmds.Abort AND NOT "R-401_DB".Status.Ready;
   IF "R-401_HMI_DB".FromHMI.Initialize THEN "R-401_HMI_DB".FromHMI.Initialize := FALSE; END_IF;
END_REGION

REGION Network 4: Start R-401
   RUNG wire#powerrail
      Contact( "R-401_HMI_DB".FromHMI.Start )
      I_Contact( "R-401_DB".Status.Aborting )
      I_Contact( "R-401_DB".Status.Initializing )
      wire#w1
      I_Contact( "R-401_DB".Status.Running )
      I_Contact( "R-401_DB".Cmds.Abort )
      Coil( "R-401_DB".Cmds.Start )
   END_RUNG
   RUNG wire#powerrail
      Contact( "R-401_DB".Cmds.Start )
   END_RUNG wire#w1
   RUNG wire#powerrail
      Contact( "R-401_HMI_DB".FromHMI.Start )
      R_Coil( "R-401_HMI_DB".FromHMI.Start )
   END_RUNG
   // the same network as SCL:
   "R-401_DB".Cmds.Start := (("R-401_HMI_DB".FromHMI.Start AND NOT "R-401_DB".Status.Aborting AND NOT "R-401_DB".Status.Initializing) OR "R-401_DB".Cmds.Start) AND NOT "R-401_DB".Status.Running AND NOT "R-401_DB".Cmds.Abort;
   IF "R-401_HMI_DB".FromHMI.Start THEN "R-401_HMI_DB".FromHMI.Start := FALSE; END_IF;
END_REGION

REGION Network 5: Procedure Selected